   "86_Times_STEP_MAX_TIME_STP_350" : Time = PLC "86_Times".STEP_MAX_TIME_STP_350, 1 s
   "86_Times_STEP_MAX_TIME_STP_230" : Time = PLC "86_Times".STEP_MAX_TIME_STP_230, 1 s
   "20_TANKS_IP_DATA_RIO_02_FIRST_TANK_GTT_ISOL_VALVE_CLSD" : Bool = PLC "20_TANKS_IP_DATA".RIO_02.FIRST_TANK.GTT_ISOL_VALVE_CLSD AT %DB1.DBW0, 1 s
   "86_Times_STEP_MAX_TIME_STP_360" : Time = PLC "86_Times".STEP_MAX_TIME_STP_360, 1 s
   "40_TANKS_OP_DATA_RIO_02_VENT_B_2P" : Bool = PLC "40_TANKS_OP_DATA".RIO_02_VENT_B_2P AT %DB1.DBW0, 1 s
   "2019_AUT_MAN_CNTRL_STBD_GTT_VLV_MAN" : Bool = PLC "2019_AUT_MAN_CNTRL".STBD_GTT_VLV_MAN AT %DB1.DBW0, 1 s
   "14_DQ_DATA_CV_422_2P" : Bool = PLC "14_DQ_DATA".CV_422_2P AT %DB1.DBW0, 1 s
   "14_DQ_DATA_CV_421_2S" : Bool = PLC "14_DQ_DATA".CV_421_2S AT %DB1.DBW0, 1 s
   "2086_Times_DEOX_PRE_GTT_OPN_DLY" : Time = PLC "2086_Times".DEOX_PRE_GTT_OPN_DLY AT %DB1.DBW0, 1 s
   "2086_Times_DEOX_PRE_GTT_CLS_DLY" : Time = PLC "2086_Times".DEOX_PRE_GTT_CLS_DLY AT %DB1.DBW0, 1 s
   "2086_Times_REOX_PRE_GTT_OPN_DLY" : Time = PLC "2086_Times".REOX_PRE_GTT_OPN_DLY AT %DB1.DBW0, 1 s
   "2086_Times_REOX_PRE_GTT_CLS_DLY" : Time = PLC "2086_Times".REOX_PRE_GTT_CLS_DLY AT %DB1.DBW0, 1 s
   "2086_Times_AT_DEOX_CNF_TIME" : Time = PLC "2086_Times".AT_DEOX_CNF_TIME AT %DB1.DBW0, 1 s
   "2086_Times_AT_REOX_CNF_TIME" : Time = PLC "2086_Times".AT_REOX_CNF_TIME AT %DB1.DBW0, 1 s
   "2084_Setpoints_FIT418_LoLo" : Real = PLC "84_Setpoints".TIT401_High AT %DB1.DBW0, 1 s
   "2084_Setpoints_PIT424_HiHi" : Real = PLC "2084_Setpoints".PIT424_HiHi AT %DB1.DBW0, 1 s
   "2084_Setpoints_PIT424_Lo" : Real = PLC "2084_Setpoints".PIT424_Lo AT %DB1.DBW0, 1 s
   "2084_Setpoints_PIT424_LoLo" : Real = PLC "2084_Setpoints".PIT424_LoLo AT %DB1.DBW0, 1 s
   "2084_Setpoints_PIT415_HiHi" : Real = PLC "2084_Setpoints".PIT415_HiHi AT %DB1.DBW0, 1 s
   "2084_Setpoints_PIT415_Hi" : Real = PLC "2084_Setpoints".PIT415_Hi AT %DB1.DBW0, 1 s
   "2084_Setpoints_PIT415_Lo" : Real = PLC "2084_Setpoints".PIT415_Lo AT %DB1.DBW0, 1 s
   "2084_Setpoints_PIT415_LoLo" : Real = PLC "2084_Setpoints".PIT415_LoLo AT %DB1.DBW0, 1 s
   "2084_Setpoints_FIT418_Lo" : Real = PLC "2084_Setpoints".FIT418_Lo AT %DB1.DBW0, 1 s
   "2084_Setpoints_FIT418_Hi" : Real = PLC "2084_Setpoints".FIT418_Hi AT %DB1.DBW0, 1 s
   "20_TANKS_IP_DATA_RIO_02_FIRST_TANK_TANK_VENT_A_CLSD" : Bool = PLC "20_TANKS_IP_DATA".RIO_02.FIRST_TANK.TANK_VENT_A_CLSD AT %DB1.DBW0, 1 s
   "2084_Setpoints_TT436_HiHi" : Real = PLC "FIT418_FPT__ALM_ANALOG_DB"."VERY HIGH LEVEL VALUE (HH)" AT %DB1.DBW0, 1 s
   "2084_Setpoints_PH_SP" : Real = PLC "2084_Setpoints".PH_SP AT %DB1.DBW0, 1 s
   "2084_Setpoints_FIT418_HiHi" : Real = PLC "2084_Setpoints".FIT418_HiHi AT %DB1.DBW0, 1 s
   "2019_AUT_MAN_CNTRL_PORT_GTT_VLV_MAN" : Bool = PLC "2019_AUT_MAN_CNTRL".PORT_GTT_VLV_MAN AT %DB1.DBW0, 1 s
   "2084_Setpoints_FIT420_LoLo" : Real = PLC "2084_Setpoints".FIT420_LoLo AT %DB1.DBW0, 1 s
   "2084_Setpoints_FIT420_Hi" : Real = PLC "2084_Setpoints".FIT420_Hi AT %DB1.DBW0, 1 s
   "2084_Setpoints_FIT420_HiHi" : Real = PLC "2084_Setpoints".FIT420_HiHi AT %DB1.DBW0, 1 s
   "2084_Setpoints_LT422_Lo" : Real = PLC "2084_Setpoints".LT422_Lo AT %DB1.DBW0, 1 s
   "2084_Setpoints_LT422_Hi" : Real = PLC "2084_Setpoints".LT422_Hi AT %DB1.DBW0, 1 s
   "2084_Setpoints_TT436_Hi" : Real = PLC "2084_Setpoints".TT436_Hi AT %DB1.DBW0, 1 s
   "2084_Setpoints_DO_SP" : Real = PLC "2084_Setpoints".DO_SP AT %DB1.DBW0, 1 s
   "2084_Setpoints_FIT420_Lo" : Real = PLC "2084_Setpoints".FIT420_Lo AT %DB1.DBW0, 1 s
   "20_TANKS_IP_DATA_RIO_02_SECOND_TANK_GTT_ISOL_VALVE_CLSD" : Bool = PLC "20_TANKS_IP_DATA".RIO_02.SECOND_TANK.GTT_ISOL_VALVE_CLSD AT %DB1.DBW0, 1 s
   "2084_Setpoints_PIT424_Hi" : Real = PLC "2084_Setpoints".PIT424_Hi AT %DB1.DBW0, 1 s
   "20_TANKS_IP_DATA_RIO_02_SECOND_TANK_DECK_IG_PRESS" : Real = PLC "20_TANKS_IP_DATA".RIO_02.SECOND_TANK.DECK_IG_PRESS AT %DB1.DBW0, 1 s
   "20_TANKS_IP_DATA_RIO_02_FIRST_TANK_TANK_VENT_B_CLSD" : Bool = PLC "20_TANKS_IP_DATA".RIO_02.FIRST_TANK.TANK_VENT_B_CLSD AT %DB1.DBW0, 1 s
   "20_TANKS_IP_DATA_RIO_02_SECOND_TANK_GTT_ISOL_VALVE_OPEN" : Bool = PLC "20_TANKS_IP_DATA".RIO_02.SECOND_TANK.GTT_ISOL_VALVE_OPEN AT %DB1.DBW0, 1 s
   "20_TANKS_IP_DATA_RIO_02_FIRST_TANK_TANK_VENT_B_OPEN" : Bool = PLC "20_TANKS_IP_DATA".RIO_02.FIRST_TANK.TANK_VENT_B_OPEN AT %DB1.DBW0, 1 s
   "40_TANKS_OP_DATA_RIO_02_VENT_B_2P(1)" : Bool = PLC "40_TANKS_OP_DATA".RIO_02_VENT_B_2P AT %DB1.DBW0, 1 s
   "20_TANKS_IP_DATA_RIO_02_SECOND_TANK_TANK_VENT_B_CLSD" : Bool = PLC "20_TANKS_IP_DATA".RIO_02.SECOND_TANK.TANK_VENT_B_CLSD AT %DB1.DBW0, 1 s
   "40_TANKS_OP_DATA_RIO_02_VENT_B_2S(1)" : Bool = PLC "40_TANKS_OP_DATA".RIO_02_VENT_B_2S AT %DB1.DBW0, 1 s
   "20_TANKS_IP_DATA_RIO_02_SECOND_TANK_TANK_VENT_A_OPEN" : Bool = PLC "20_TANKS_IP_DATA".RIO_02.SECOND_TANK.TANK_VENT_A_OPEN AT %DB1.DBW0, 1 s
   "20_TANKS_IP_DATA_RIO_02_SECOND_TANK_TANK_VENT_A_CLSD" : Bool = PLC "20_TANKS_IP_DATA".RIO_02.SECOND_TANK.TANK_VENT_A_CLSD AT %DB1.DBW0, 1 s
   "20_TANKS_IP_DATA_RIO_02_FIRST_TANK_BWT_LEVEL_HIHI" : Bool = PLC "20_TANKS_IP_DATA".RIO_02.FIRST_TANK.BWT_LEVEL_HIHI AT %DB1.DBW0, 1 s
   "20_TANKS_IP_DATA_RIO_02_SECOND_TANK_BWT_LEVEL_HIHI" : Bool = PLC "20_TANKS_IP_DATA".RIO_02.SECOND_TANK.BWT_LEVEL_HIHI AT %DB1.DBW0, 1 s
   "20_TANKS_IP_DATA_RIO_02_SECOND_TANK_TANK_VENT_B_OPEN" : Bool = PLC "20_TANKS_IP_DATA".RIO_02.SECOND_TANK.TANK_VENT_B_OPEN AT %DB1.DBW0, 1 s
   "20_TANKS_IP_DATA_RIO_02_SECOND_TANK_TANKS_PRESS_HIHI" : Bool = PLC "20_TANKS_IP_DATA".RIO_02.SECOND_TANK.TANKS_PRESS_HIHI AT %DB1.DBW0, 1 s
   "20_TANKS_IP_DATA_RIO_02_SECOND_TANK_MBG_FLOW" : Real = PLC "20_TANKS_IP_DATA".RIO_02.SECOND_TANK.MBG_FLOW AT %DB1.DBW0, 1 s
   "20_TANKS_IP_DATA_RIO_02_FIRST_TANK_TANKS_PRESS" : Real = PLC "20_TANKS_IP_DATA".RIO_02.FIRST_TANK.TANKS_PRESS AT %DB1.DBW0, 1 s
   "20_TANKS_IP_DATA_RIO_02_FIRST_TANK_USD_FLOW" : Real = PLC "20_TANKS_IP_DATA".RIO_02.FIRST_TANK.USD_FLOW AT %DB1.DBW0, 1 s
   "20_TANKS_IP_DATA_RIO_02_FIRST_TANK_TANKS_PRESS_HIHI" : Bool = PLC "20_TANKS_IP_DATA".RIO_02.FIRST_TANK.TANKS_PRESS_HIHI AT %DB1.DBW0, 1 s
   "20_TANKS_IP_DATA_RIO_02_FIRST_TANK_MBG_FLOW" : Real = PLC "20_TANKS_IP_DATA".RIO_02.FIRST_TANK.MBG_FLOW AT %DB1.DBW0, 1 s
   "20_TANKS_IP_DATA_RIO_02_FIRST_TANK_O2_MONITOR" : Real = PLC "20_TANKS_IP_DATA".RIO_02.FIRST_TANK.O2_MONITOR AT %DB1.DBW0, 1 s
   "20_TANKS_IP_DATA_RIO_02_SECOND_TANK_USD_FLOW" : Real = PLC "20_TANKS_IP_DATA".RIO_02.SECOND_TANK.USD_FLOW AT %DB1.DBW0, 1 s
   "20_TANKS_IP_DATA_RIO_02_SECOND_TANK_TANKS_PRESS" : Real = PLC "20_TANKS_IP_DATA".RIO_02.SECOND_TANK.TANKS_PRESS AT %DB1.DBW0, 1 s
   "20_TANKS_IP_DATA_RIO_02_SECOND_TANK_O2_MONITOR" : Real = PLC "20_TANKS_IP_DATA".RIO_02.SECOND_TANK.O2_MONITOR AT %DB1.DBW0, 1 s
   "62_Warning_Data_GCU_WARNING_WORD_09(1)" : Word = PLC "62_Warning_Data".GCU_WARNING_WORD_09 AT %DB62.DBW16, 1 s
   "62_Warning_Data_GCU_WARNING_WORD_01(1)" : Word = PLC "62_Warning_Data".GCU_WARNING_WORD_01 AT %DB62.DBW0, 1 s
   "62_Warning_Data_BWTS_WARNING_WORD_10" : Word = PLC "62_Warning_Data".BWTS_WARNING_WORD_10 AT %DB62.DBW18, 1 s
   "62_Warning_Data_BWTS_WARNING_WORD_11" : Word = PLC "62_Warning_Data".BWTS_WARNING_WORD_11 AT %DB62.DBW20, 1 s
   "62_Warning_Data_GCU_WARNING_WORD_02(1)" : Word = PLC "62_Warning_Data".GCU_WARNING_WORD_02 AT %DB62.DBW2, 1 s
   "62_Warning_Data_GCU_WARNING_WORD_03(1)" : Word = PLC "62_Warning_Data".GCU_WARNING_WORD_03 AT %DB62.DBW4, 1 s
   "62_Warning_Data_GCU_WARNING_WORD_04(1)" : Word = PLC "62_Warning_Data".GCU_WARNING_WORD_04 AT %DB62.DBW6, 1 s
   "62_Warning_Data_GCU_WARNING_WORD_05(1)" : Word = PLC "62_Warning_Data".GCU_WARNING_WORD_05 AT %DB62.DBW8, 1 s
   "62_Warning_Data_GCU_WARNING_WORD_06(1)" : Word = PLC "62_Warning_Data".GCU_WARNING_WORD_06 AT %DB62.DBW10, 1 s
   "62_Warning_Data_GCU_WARNING_WORD_07(1)" : Word = PLC "62_Warning_Data".GCU_WARNING_WORD_07 AT %DB62.DBW12, 1 s
   "62_Warning_Data_GCU_WARNING_WORD_08(1)" : Word = PLC "62_Warning_Data".GCU_WARNING_WORD_08 AT %DB62.DBW14, 1 s
   "Record Data Tag" : Int AT %DB1.DBX0.0
   "Recipe Tag" : Int, internal
   "Data_From_WBT_Level_APT" : Real = PLC Data_From_WBT.Level_APT, 1 s
   "Data_From_WBT_Level_WBT_6P" : Real = PLC Data_From_WBT.Level_WBT_6P, 1 s
   "Data_From_WBT_Level_WBT_5P" : Real = PLC Data_From_WBT.Level_WBT_5P, 1 s
   "Data_From_WBT_Level_WBT_4P" : Real = PLC Data_From_WBT.Level_WBT_4P, 1 s
   "Data_From_WBT_Level_WBT_3P" : Real = PLC Data_From_WBT.Level_WBT_3P, 1 s
   "Data_From_WBT_Level_WBT_2P" : Real = PLC Data_From_WBT.Level_WBT_2P, 1 s
   "Data_From_WBT_Level_WBT_1P" : Real = PLC Data_From_WBT.Level_WBT_1P, 1 s
   "Data_From_WBT_Level_FPT" : Real = PLC Data_From_WBT.Level_FPT, 1 s
   "Data_From_WBT_Level_WBT_1S" : Real = PLC Data_From_WBT.Level_WBT_1S, 1 s
   "Data_From_WBT_Level_WBT_2S" : Real = PLC Data_From_WBT.Level_WBT_2S, 1 s
   "Data_From_WBT_Level_WBT_3S" : Real = PLC Data_From_WBT.Level_WBT_3S, 1 s
   "Data_From_WBT_Level_WBT_4S" : Real = PLC Data_From_WBT.Level_WBT_4S, 1 s
   "Data_From_WBT_Level_WBT_5S" : Real = PLC Data_From_WBT.Level_WBT_5S, 1 s
   "Data_From_WBT_Level_WBT_6S" : Real = PLC Data_From_WBT.Level_WBT_6S, 1 s
   "Data_From_WBT_Level_APT(1)" : Real = PLC Data_From_WBT.Level_APT, 1 s
   "Data_From_WBT_Level_APT m" : Real = PLC Data_From_WBT."Level_APT m", 1 s
   "Data_From_WBT_Level_WBT_6S m" : Real = PLC Data_From_WBT."Level_WBT_6S m", 1 s
   "Data_From_WBT_Level_WBT_5S m" : Real = PLC Data_From_WBT."Level_WBT_5S m", 1 s
   "Data_From_WBT_Level_WBT_4S m" : Real = PLC Data_From_WBT."Level_WBT_4S m", 1 s
   "Data_From_WBT_Level_WBT_3S m" : Real = PLC Data_From_WBT."Level_WBT_3S m", 1 s
   "Data_From_WBT_Level_WBT_2S m" : Real = PLC Data_From_WBT."Level_WBT_2S m", 1 s
   "Data_From_WBT_Level_WBT_1S m" : Real = PLC Data_From_WBT."Level_WBT_1S m", 1 s
   "Data_From_WBT_Level_FPT m" : Real = PLC Data_From_WBT."Level_FPT m", 1 s
   "Data_From_WBT_Level_WBT_1P m" : Real = PLC Data_From_WBT."Level_WBT_1P m", 1 s
   "Data_From_WBT_Level_WBT_2P m" : Real = PLC Data_From_WBT."Level_WBT_2P m", 1 s
   "Data_From_WBT_Level_WBT_3P m" : Real = PLC Data_From_WBT."Level_WBT_3P m", 1 s
   "Data_From_WBT_Level_WBT_4P m" : Real = PLC Data_From_WBT."Level_WBT_4P m", 1 s
   "Data_From_WBT_Level_WBT_5P m" : Real = PLC Data_From_WBT."Level_WBT_5P m", 1 s
   "Data_From_WBT_Level_WBT_6P m" : Real = PLC Data_From_WBT."Level_WBT_6P m", 1 s
   "HEART BEAT TRUE" : Bool = PLC "68_Sys_Status_Data"."TRUE for HMI" AT %M1.2, 100 ms
   "Warn To Start IGG" : Bool = PLC "82_To_HMI"."Warn to Start IGG", 1 s
      on ChangeValue: "TimeRemainingToTreatment"()

discrete alarms
   129: 'PIT-359 - HIGH HIGH', class IGG Alarms, trigger "Alarms_Acknowledge_IGG_ALARM_ACKNLG_2" bit 1
   130: 'PIT-316 - HIGH HIGH', class IGG Alarms, trigger "Alarms_Acknowledge_IGG_ALARM_ACKNLG_2" bit 3
   131: 'PIT-359 - LOW LOW', class IGG Alarms, trigger "Alarms_Acknowledge_IGG_ALARM_ACKNLG_2" bit 0
   132: 'PIT-316 - LOW LOW', class IGG Alarms, trigger "Alarms_Acknowledge_IGG_ALARM_ACKNLG_2" bit 2
   279: 'IGG_MESSAGE_WORD_02_BIT_14', class IGG Messages, trigger "64_Message_Data_IGG_MESSAGE_WORD_02" bit 6
   133: 'PIT-359 - HIGH HIGH', class IGG Alarms, trigger "Alarms_Acknowledge_IGG_ALARM_ACKNLG_2" bit 4
   134: 'TIT-401 - HIGH HIGH', class IGG Alarms, trigger "Alarms_Acknowledge_IGG_ALARM_ACKNLG_2" bit 10
   135: 'PIT-102 CA PRESSURE - FAULT', class IGG Alarms, trigger "Alarms_Acknowledge_IGG_ALARM_ACKNLG_2" bit 9
   136: 'PIT-402 IG OUTLET PRESSURE - HIGH HIGH', class IGG Alarms, trigger "Alarms_Acknowledge_IGG_ALARM_ACKNLG_2" bit 12
   137: 'PIT-402 IG OUTLET PRESSURE - LOW LOW', class IGG Alarms, trigger "Alarms_Acknowledge_IGG_ALARM_ACKNLG_2" bit 11
   138: 'IGG_ALARM_WORD_02_BIT_14', class IGG Alarms, trigger "Alarms_Acknowledge_IGG_ALARM_ACKNLG_2" bit 6
   139: 'IGG_ALARM_WORD_02_BIT_13', class IGG Alarms, trigger "Alarms_Acknowledge_IGG_ALARM_ACKNLG_2" bit 5
   140: 'PIT-102 CA PRESSURE - LOW LOW', class IGG Alarms, trigger "Alarms_Acknowledge_IGG_ALARM_ACKNLG_2" bit 8
   141: 'IGG_ALARM_WORD_02_BIT_15', class IGG Alarms, trigger "Alarms_Acknowledge_IGG_ALARM_ACKNLG_2" bit 7
   142: 'EMERGENCY STOP ACTIVE', class IGG Alarms, trigger "Alarms_Acknowledge_IGG_ALARM_ACKNLG_1" bit 15
   143: 'ATMOSPHERIC O2 SENSOR 1 - LOW LOW', class IGG Alarms, trigger "Alarms_Acknowledge_IGG_ALARM_ACKNLG_1" bit 1
   144: 'BC ALARM ACTIVE', class IGG Alarms, trigger "Alarms_Acknowledge_IGG_ALARM_ACKNLG_1" bit 0
   145: 'ATMOSPHERIC O2 SENSOR 2 - LOW LOW', class IGG Alarms, trigger "Alarms_Acknowledge_IGG_ALARM_ACKNLG_1" bit 2
   146: 'E-500B FUEL PUMP - NOT RUNNING', class IGG Alarms, trigger "Alarms_Acknowledge_IGG_ALARM_ACKNLG_1" bit 4
   147: 'E-500A FUEL PUMP - NOT RUNNING', class IGG Alarms, trigger "Alarms_Acknowledge_IGG_ALARM_ACKNLG_1" bit 3
   383: 'BC_EVENT_WORD_02_BIT_6', class BC Events, trigger "66_Event_Data_BC_EVENT_WORD_02" bit 14
   382: 'BC_EVENT_WORD_02_BIT_5', class BC Events, trigger "66_Event_Data_BC_EVENT_WORD_02" bit 13
   384: 'BC_EVENT_WORD_02_BIT_7', class BC Events, trigger "66_Event_Data_BC_EVENT_WORD_02" bit 15
   278: 'IGG_MESSAGE_WORD_02_BIT_13', class IGG Messages, trigger "64_Message_Data_IGG_MESSAGE_WORD_02" bit 5
   277: 'IGG_MESSAGE_WORD_02_BIT_12', class IGG Messages, trigger "64_Message_Data_IGG_MESSAGE_WORD_02" bit 4
   148: 'P-301 CSW PUMP - TRIPPED', class IGG Alarms, trigger "Alarms_Acknowledge_IGG_ALARM_ACKNLG_1" bit 11
   149: 'IGG AUTO INTERLOCKS NOT OK', class IGG Alarms, trigger "Alarms_Acknowledge_IGG_ALARM_ACKNLG_1" bit 10
   150: 'E-500A FUEL PUMP - TRIPPED', class IGG Alarms, trigger "Alarms_Acknowledge_IGG_ALARM_ACKNLG_1" bit 12
   151: 'E-139 CAB INVERTER - FAULT', class IGG Alarms, trigger "Alarms_Acknowledge_IGG_ALARM_ACKNLG_1" bit 14
   152: 'E-500B FUEL PUMP - TRIPPED', class IGG Alarms, trigger "Alarms_Acknowledge_IGG_ALARM_ACKNLG_1" bit 13
   153: 'IGG_ALARM_WORD_01_BIT_14', class IGG Alarms, trigger "Alarms_Acknowledge_IGG_ALARM_ACKNLG_1" bit 6
   154: 'E-139 CAB NOT READY3', class IGG Alarms, trigger "Alarms_Acknowledge_IGG_ALARM_ACKNLG_1" bit 5
   155: 'IGG_ALARM_WORD_01_BIT_15', class IGG Alarms, trigger "Alarms_Acknowledge_IGG_ALARM_ACKNLG_1" bit 7
   156: 'SLAVE PLC HEART BEAT MISSING', class IGG Alarms, trigger "Alarms_Acknowledge_IGG_ALARM_ACKNLG_1" bit 9
   157: 'MASTER PLC HEART BEAT MISSING', class IGG Alarms, trigger "Alarms_Acknowledge_IGG_ALARM_ACKNLG_1" bit 8
   158: 'PIT-402 IG PRESSURE - OUT OF RANGE', class IGG Alarms, trigger "Alarms_Acknowledge_IGG_ALARM_ACKNLG_2" bit 13
   55: 'IGG_ALARM_WORD_04_BIT_14', class IGG Alarms, trigger "Alarms_Acknowledge_IGG_ALARM_ACKNLG_4" bit 6
   54: 'CORRECT PHASE ROTATION - FAULT', class IGG Alarms, trigger "Alarms_Acknowledge_IGG_ALARM_ACKNLG_4" bit 5
   56: 'IGG_ALARM_WORD_04_BIT_15', class IGG Alarms, trigger "Alarms_Acknowledge_IGG_ALARM_ACKNLG_4" bit 7
   58: 'CV-312 - FAULT', class IGG Alarms, trigger "Alarms_Acknowledge_IGG_ALARM_ACKNLG_4" bit 9
   57: 'CV-311 - FAULT', class IGG Alarms, trigger "Alarms_Acknowledge_IGG_ALARM_ACKNLG_4" bit 8
   50: 'TIT-319 INLET CSW TEMP - FAULT AND TIT-401 AND TIT-360 - FAULT', class IGG Alarms, trigger "Alarms_Acknowledge_IGG_ALARM_ACKNLG_4" bit 1
   49: 'TIT-319 INLET CSW TEMP - FAULT AND TS-006 - FAULT', class IGG Alarms, trigger "Alarms_Acknowledge_IGG_ALARM_ACKNLG_4" bit 0
   51: 'TIT-360 OUTLET CSW TEMP - HIGH HIGH0', class IGG Alarms, trigger "Alarms_Acknowledge_IGG_ALARM_ACKNLG_4" bit 2
   53: 'E-139 NOT RUNNING2', class IGG Alarms, trigger "Alarms_Acknowledge_IGG_ALARM_ACKNLG_4" bit 4
   52: 'TIT-360 OUTLET CSW TEMP - HIGH HIGH AND TIT-401 - FAULT', class IGG Alarms, trigger "Alarms_Acknowledge_IGG_ALARM_ACKNLG_4" bit 3
   59: 'CV-321 - FAULT', class IGG Alarms, trigger "Alarms_Acknowledge_IGG_ALARM_ACKNLG_4" bit 10
   65: 'IGG ALARM ACTIVE', class BC Alarms, trigger "BC_ALARM_ACKNLG_1" bit 0
   282: 'IGG_MESSAGE_WORD_02_BIT_1', class IGG Messages, trigger "64_Message_Data_IGG_MESSAGE_WORD_02" bit 9
   66: 'PS-101 PRESSURE NOT PRESENT - FAULT', class BC Alarms, trigger "BC_ALARM_ACKNLG_1" bit 1
   69: 'FD-001 FLAME SIGNAL - OUT OF RANGE', class BC Alarms, trigger "BC_ALARM_ACKNLG_1" bit 4
   68: 'O2 SYSTEM POWER NOT HEALTHY', class BC Alarms, trigger "BC_ALARM_ACKNLG_1" bit 3
   61: 'CV-401 - FAULT', class IGG Alarms, trigger "Alarms_Acknowledge_IGG_ALARM_ACKNLG_4" bit 12
   60: 'CV-322 - FAULT', class IGG Alarms, trigger "Alarms_Acknowledge_IGG_ALARM_ACKNLG_4" bit 11
   62: 'CV-431 - FAULT', class IGG Alarms, trigger "Alarms_Acknowledge_IGG_ALARM_ACKNLG_4" bit 13
   64: 'SAFETY SYSTEM INTERLOCK', class IGG Alarms, trigger "Alarms_Acknowledge_IGG_ALARM_ACKNLG_4" bit 15
   63: 'CV-432 - FAULT', class IGG Alarms, trigger "Alarms_Acknowledge_IGG_ALARM_ACKNLG_4" bit 14
   35: 'TIT-315 SHELL CSW TEMP - HIGH HIGH AND TIT-401 - FAULT', class IGG Alarms, trigger "Alarms_Acknowledge_IGG_ALARM_ACKNLG_3" bit 2
   34: 'TIT-315 SHELL CSW TEMP - HIGH HIGH AND TS-006 - FAULT', class IGG Alarms, trigger "Alarms_Acknowledge_IGG_ALARM_ACKNLG_3" bit 1
   36: 'PIT-316 OUTLET CSW PRESSURE AND FS-317 - FAULT', class IGG Alarms, trigger "Alarms_Acknowledge_IGG_ALARM_ACKNLG_3" bit 3
   38: 'PIT-316 OUTLET CSW PRESSURE AND TS-006 - FAULT', class IGG Alarms, trigger "Alarms_Acknowledge_IGG_ALARM_ACKNLG_3" bit 5
   37: 'PIT-316 OUTLET CSW PRESSURE AND TIT-315 - FAULT', class IGG Alarms, trigger "Alarms_Acknowledge_IGG_ALARM_ACKNLG_3" bit 4
   159: 'TIT-360 - HIGH HIGH', class IGG Alarms, trigger "Alarms_Acknowledge_IGG_ALARM_ACKNLG_2" bit 15
   160: 'TIT-319 - HIGH HIGH', class IGG Alarms, trigger "Alarms_Acknowledge_IGG_ALARM_ACKNLG_2" bit 14
   280: 'IGG_MESSAGE_WORD_02_BIT_15', class IGG Messages, trigger "64_Message_Data_IGG_MESSAGE_WORD_02" bit 7
   33: 'TIT-315 SHELL CSW TEMP - HIGH HIGH AND FS-317 - FAULT', class IGG Alarms, trigger "Alarms_Acknowledge_IGG_ALARM_ACKNLG_3" bit 0
   70: 'E-600 O2 ANALYSER CONTENT - OUT OF RANGE', class BC Alarms, trigger "BC_ALARM_ACKNLG_1" bit 5
   39: 'IGG_ALARM_WORD_03_BIT_14', class IGG Alarms, trigger "Alarms_Acknowledge_IGG_ALARM_ACKNLG_3" bit 6
   46: 'TIT-401 IG TEMP - HIGH HIGH AND TIT-360 - FAULT', class IGG Alarms, trigger "Alarms_Acknowledge_IGG_ALARM_ACKNLG_3" bit 13
   45: 'TIT-401 IG TEMP - HIGH HIGH AND TS-403 - FAULT', class IGG Alarms, trigger "Alarms_Acknowledge_IGG_ALARM_ACKNLG_3" bit 12
   47: 'IGG_ALARM_WORD_03_BIT_6', class IGG Alarms, trigger "Alarms_Acknowledge_IGG_ALARM_ACKNLG_3" bit 14
   281: 'IGG_MESSAGE_WORD_02_BIT_0', class IGG Messages, trigger "64_Message_Data_IGG_MESSAGE_WORD_02" bit 8
   48: 'IGG_ALARM_WORD_03_BIT_7', class IGG Alarms, trigger "Alarms_Acknowledge_IGG_ALARM_ACKNLG_3" bit 15
   41: 'PIT-112/113 TIER ALARM - PRESSURE NOT OK', class IGG Alarms, trigger "Alarms_Acknowledge_IGG_ALARM_ACKNLG_3" bit 8
   40: 'IGG_ALARM_WORD_03_BIT_15', class IGG Alarms, trigger "Alarms_Acknowledge_IGG_ALARM_ACKNLG_3" bit 7
   42: 'PIT-102 CA PRESSURE - LOW LOW AND FDU - FAULT', class IGG Alarms, trigger "Alarms_Acknowledge_IGG_ALARM_ACKNLG_3" bit 9
   44: 'IGG ALARM WORD', class IGG Alarms, trigger "Alarms_Acknowledge_IGG_ALARM_ACKNLG_3" bit 11
   43: 'PIT-102 CA PRESSURE - LOW LOW AND PIT-402 - FAULT', class IGG Alarms, trigger "Alarms_Acknowledge_IGG_ALARM_ACKNLG_3" bit 10
   381: 'BC_EVENT_WORD_02_BIT_4', class BC Events, trigger "66_Event_Data_BC_EVENT_WORD_02" bit 12
   330: 'IGG_EVENT_WORD_01_BIT_1', class IGG Events, trigger "66_Event_Data_IGG_EVENT_WORD_01" bit 9
   329: 'IGG_EVENT_WORD_01_BIT_0', class IGG Events, trigger "66_Event_Data_IGG_EVENT_WORD_01" bit 8
   331: 'IGG_EVENT_WORD_01_BIT_2', class IGG Events, trigger "66_Event_Data_IGG_EVENT_WORD_01" bit 10
   333: 'IGG_EVENT_WORD_01_BIT_4', class IGG Events, trigger "66_Event_Data_IGG_EVENT_WORD_01" bit 12
   332: 'IGG_EVENT_WORD_01_BIT_3', class IGG Events, trigger "66_Event_Data_IGG_EVENT_WORD_01" bit 11
   325: 'IGG_EVENT_WORD_01_BIT_12', class IGG Events, trigger "66_Event_Data_IGG_EVENT_WORD_01" bit 4
   324: 'IGG_EVENT_WORD_01_BIT_11', class IGG Events, trigger "66_Event_Data_IGG_EVENT_WORD_01" bit 3
   326: 'IGG_EVENT_WORD_01_BIT_13', class IGG Events, trigger "66_Event_Data_IGG_EVENT_WORD_01" bit 5
   328: 'IGG_EVENT_WORD_01_BIT_15', class IGG Events, trigger "66_Event_Data_IGG_EVENT_WORD_01" bit 7
   327: 'IGG_EVENT_WORD_01_BIT_14', class IGG Events, trigger "66_Event_Data_IGG_EVENT_WORD_01" bit 6
   338: 'IGG_EVENT_WORD_02_BIT_9', class IGG Events, trigger "66_Event_Data_IGG_EVENT_WORD_02" bit 1
   337: 'IGG_EVENT_WORD_02_BIT_8', class IGG Events, trigger "66_Event_Data_IGG_EVENT_WORD_02" bit 0
   339: 'IGG_EVENT_WORD_02_BIT_10', class IGG Events, trigger "66_Event_Data_IGG_EVENT_WORD_02" bit 2
   341: 'IGG_EVENT_WORD_02_BIT_12', class IGG Events, trigger "66_Event_Data_IGG_EVENT_WORD_02" bit 4
   340: 'IGG_EVENT_WORD_02_BIT_11', class IGG Events, trigger "66_Event_Data_IGG_EVENT_WORD_02" bit 3
   335: 'IGG_EVENT_WORD_01_BIT_6', class IGG Events, trigger "66_Event_Data_IGG_EVENT_WORD_01" bit 14
   334: 'IGG_EVENT_WORD_01_BIT_5', class IGG Events, trigger "66_Event_Data_IGG_EVENT_WORD_01" bit 13
   336: 'IGG_EVENT_WORD_01_BIT_7', class IGG Events, trigger "66_Event_Data_IGG_EVENT_WORD_01" bit 15
   276: 'IGG_MESSAGE_WORD_02_BIT_11', class IGG Messages, trigger "64_Message_Data_IGG_MESSAGE_WORD_02" bit 3
   259: 'IGG_MESSAGE_WORD_01_BIT_10', class IGG Messages, trigger "64_Message_Data_IGG_MESSAGE_WORD_01" bit 2
   267: 'IGG_MESSAGE_WORD_01_BIT_2', class IGG Messages, trigger "64_Message_Data_IGG_MESSAGE_WORD_01" bit 10
   268: 'IGG_MESSAGE_WORD_01_BIT_3', class IGG Messages, trigger "64_Message_Data_IGG_MESSAGE_WORD_01" bit 11
   273: 'IGG_MESSAGE_WORD_02_BIT_8', class IGG Messages, trigger "64_Message_Data_IGG_MESSAGE_WORD_02" bit 0
   265: 'IGG_MESSAGE_WORD_01_BIT_0', class IGG Messages, trigger "64_Message_Data_IGG_MESSAGE_WORD_01" bit 8
   266: 'IGG_MESSAGE_WORD_01_BIT_1', class IGG Messages, trigger "64_Message_Data_IGG_MESSAGE_WORD_01" bit 9
   272: 'IGG_MESSAGE_WORD_01_BIT_7', class IGG Messages, trigger "64_Message_Data_IGG_MESSAGE_WORD_01" bit 15
   67: 'E-600 O2 ANALYSER SYSTEM - FAIL', class BC Alarms, trigger "BC_ALARM_ACKNLG_1" bit 2
   271: 'IGG_MESSAGE_WORD_01_BIT_6', class IGG Messages, trigger "64_Message_Data_IGG_MESSAGE_WORD_01" bit 14
   269: 'IGG_MESSAGE_WORD_01_BIT_4', class IGG Messages, trigger "64_Message_Data_IGG_MESSAGE_WORD_01" bit 12
   270: 'IGG_MESSAGE_WORD_01_BIT_5', class IGG Messages, trigger "64_Message_Data_IGG_MESSAGE_WORD_01" bit 13
   260: 'IGG_MESSAGE_WORD_01_BIT_11', class IGG Messages, trigger "64_Message_Data_IGG_MESSAGE_WORD_01" bit 3
   275: 'IGG_MESSAGE_WORD_02_BIT_10', class IGG Messages, trigger "64_Message_Data_IGG_MESSAGE_WORD_02" bit 2
   321: 'IGG_EVENT_WORD_01_BIT_8', class IGG Events, trigger "66_Event_Data_IGG_EVENT_WORD_01" bit 0
   323: 'IGG_EVENT_WORD_01_BIT_10', class IGG Events, trigger "66_Event_Data_IGG_EVENT_WORD_01" bit 2
   322: 'IGG_EVENT_WORD_01_BIT_9', class IGG Events, trigger "66_Event_Data_IGG_EVENT_WORD_01" bit 1
   264: 'IGG_MESSAGE_WORD_01_BIT_15', class IGG Messages, trigger "64_Message_Data_IGG_MESSAGE_WORD_01" bit 7
   274: 'IGG_MESSAGE_WORD_02_BIT_9', class IGG Messages, trigger "64_Message_Data_IGG_MESSAGE_WORD_02" bit 1
   263: 'IGG_MESSAGE_WORD_01_BIT_14', class IGG Messages, trigger "64_Message_Data_IGG_MESSAGE_WORD_01" bit 6
   261: 'IGG_MESSAGE_WORD_01_BIT_12', class IGG Messages, trigger "64_Message_Data_IGG_MESSAGE_WORD_01" bit 4
   262: 'IGG_MESSAGE_WORD_01_BIT_13', class IGG Messages, trigger "64_Message_Data_IGG_MESSAGE_WORD_01" bit 5
   342: 'IGG_EVENT_WORD_02_BIT_13', class IGG Events, trigger "66_Event_Data_IGG_EVENT_WORD_02" bit 5
   367: 'BC_EVENT_WORD_01_BIT_6', class BC Events, trigger "66_Event_Data_BC_EVENT_WORD_01" bit 14
   366: 'BC_EVENT_WORD_01_BIT_5', class BC Events, trigger "66_Event_Data_BC_EVENT_WORD_01" bit 13
   368: 'BC_EVENT_WORD_01_BIT_7', class BC Events, trigger "66_Event_Data_BC_EVENT_WORD_01" bit 15
   370: 'BC_EVENT_WORD_02_BIT_9', class BC Events, trigger "66_Event_Data_BC_EVENT_WORD_02" bit 1
   369: 'BC_EVENT_WORD_02_BIT_8', class BC Events, trigger "66_Event_Data_BC_EVENT_WORD_02" bit 0
   362: 'BC_EVENT_WORD_01_BIT_1', class BC Events, trigger "66_Event_Data_BC_EVENT_WORD_01" bit 9
   361: 'BC_EVENT_WORD_01_BIT_0', class BC Events, trigger "66_Event_Data_BC_EVENT_WORD_01" bit 8
   363: 'BC_EVENT_WORD_01_BIT_2', class BC Events, trigger "66_Event_Data_BC_EVENT_WORD_01" bit 10
   365: 'BC_EVENT_WORD_01_BIT_4', class BC Events, trigger "66_Event_Data_BC_EVENT_WORD_01" bit 12
   364: 'BC_EVENT_WORD_01_BIT_3', class BC Events, trigger "66_Event_Data_BC_EVENT_WORD_01" bit 11
   377: 'BC_EVENT_WORD_02_BIT_0', class BC Events, trigger "66_Event_Data_BC_EVENT_WORD_02" bit 8
   376: 'BC_EVENT_WORD_02_BIT_15', class BC Events, trigger "66_Event_Data_BC_EVENT_WORD_02" bit 7
   378: 'BC_EVENT_WORD_02_BIT_1', class BC Events, trigger "66_Event_Data_BC_EVENT_WORD_02" bit 9
   380: 'BC_EVENT_WORD_02_BIT_3', class BC Events, trigger "66_Event_Data_BC_EVENT_WORD_02" bit 11
   379: 'BC_EVENT_WORD_02_BIT_2', class BC Events, trigger "66_Event_Data_BC_EVENT_WORD_02" bit 10
   372: 'BC_EVENT_WORD_02_BIT_11', class BC Events, trigger "66_Event_Data_BC_EVENT_WORD_02" bit 3
   371: 'BC_EVENT_WORD_02_BIT_10', class BC Events, trigger "66_Event_Data_BC_EVENT_WORD_02" bit 2
   373: 'BC_EVENT_WORD_02_BIT_12', class BC Events, trigger "66_Event_Data_BC_EVENT_WORD_02" bit 4
   375: 'BC_EVENT_WORD_02_BIT_14', class BC Events, trigger "66_Event_Data_BC_EVENT_WORD_02" bit 6
   374: 'BC_EVENT_WORD_02_BIT_13', class BC Events, trigger "66_Event_Data_BC_EVENT_WORD_02" bit 5
   349: 'IGG_EVENT_WORD_02_BIT_4', class IGG Events, trigger "66_Event_Data_IGG_EVENT_WORD_02" bit 12
   348: 'IGG_EVENT_WORD_02_BIT_3', class IGG Events, trigger "66_Event_Data_IGG_EVENT_WORD_02" bit 11
   350: 'IGG_EVENT_WORD_02_BIT_5', class IGG Events, trigger "66_Event_Data_IGG_EVENT_WORD_02" bit 13
   352: 'IGG_EVENT_WORD_02_BIT_7', class IGG Events, trigger "66_Event_Data_IGG_EVENT_WORD_02" bit 15
   351: 'IGG_EVENT_WORD_02_BIT_6', class IGG Events, trigger "66_Event_Data_IGG_EVENT_WORD_02" bit 14
   344: 'IGG_EVENT_WORD_02_BIT_15', class IGG Events, trigger "66_Event_Data_IGG_EVENT_WORD_02" bit 7
   343: 'IGG_EVENT_WORD_02_BIT_14', class IGG Events, trigger "66_Event_Data_IGG_EVENT_WORD_02" bit 6
   345: 'IGG_EVENT_WORD_02_BIT_0', class IGG Events, trigger "66_Event_Data_IGG_EVENT_WORD_02" bit 8
   347: 'IGG_EVENT_WORD_02_BIT_2', class IGG Events, trigger "66_Event_Data_IGG_EVENT_WORD_02" bit 10
   346: 'IGG_EVENT_WORD_02_BIT_1', class IGG Events, trigger "66_Event_Data_IGG_EVENT_WORD_02" bit 9
   357: 'BC_EVENT_WORD_01_BIT_12', class BC Events, trigger "66_Event_Data_BC_EVENT_WORD_01" bit 4
   356: 'BC_EVENT_WORD_01_BIT_11', class BC Events, trigger "66_Event_Data_BC_EVENT_WORD_01" bit 3
   358: 'BC_EVENT_WORD_01_BIT_13', class BC Events, trigger "66_Event_Data_BC_EVENT_WORD_01" bit 5
   360: 'BC_EVENT_WORD_01_BIT_15', class BC Events, trigger "66_Event_Data_BC_EVENT_WORD_01" bit 7
   359: 'BC_EVENT_WORD_01_BIT_14', class BC Events, trigger "66_Event_Data_BC_EVENT_WORD_01" bit 6
   257: 'IGG_MESSAGE_WORD_01_BIT_8', class IGG Messages, trigger "64_Message_Data_IGG_MESSAGE_WORD_01" bit 0
   258: 'IGG_MESSAGE_WORD_01_BIT_9', class IGG Messages, trigger "64_Message_Data_IGG_MESSAGE_WORD_01" bit 1
   353: 'BC_EVENT_WORD_01_BIT_8', class BC Events, trigger "66_Event_Data_BC_EVENT_WORD_01" bit 0
   355: 'BC_EVENT_WORD_01_BIT_10', class BC Events, trigger "66_Event_Data_BC_EVENT_WORD_01" bit 2
   354: 'BC_EVENT_WORD_01_BIT_9', class BC Events, trigger "66_Event_Data_BC_EVENT_WORD_01" bit 1
   114: 'P-305 FRESH WATER PUMP - TRIPPED', class BC Alarms, trigger "BC_ALARM_ACKNLG_4" bit 1
   113: 'LS-001 IGG QUENCH CHAMBER LEVEL - HIGH', class BC Alarms, trigger "BC_ALARM_ACKNLG_4" bit 0
   116: 'BC_ALARM_WORD_04_BIT_11', class BC Alarms, trigger "BC_ALARM_ACKNLG_4" bit 3
   115: 'BC_ALARM_WORD_04_BIT_10', class BC Alarms, trigger "BC_ALARM_ACKNLG_4" bit 2
   284: 'IGG_MESSAGE_WORD_02_BIT_3', class IGG Messages, trigger "64_Message_Data_IGG_MESSAGE_WORD_02" bit 11
   112: 'BC_ALARM_WORD_3_BIT_15', class BC Alarms, trigger "BC_ALARM_ACKNLG_3" bit 15
   315: 'BC_MESSAGE_WORD_02_BIT_2', class BC Messages, trigger "64_Message_Data_BC_MESSAGE_WORD_02" bit 10
   316: 'BC_MESSAGE_WORD_02_BIT_3', class BC Messages, trigger "64_Message_Data_BC_MESSAGE_WORD_02" bit 11
   122: 'TS-006 IG SHELL TEMP HI SWITCH AND TIT-360 - FAULT', class BC Alarms, trigger "BC_ALARM_ACKNLG_4" bit 9
   121: 'TS-006 IGG SHELL TEMPERATURE - HIGH', class BC Alarms, trigger "BC_ALARM_ACKNLG_4" bit 8
   124: 'TS-403 IG TEMP - HIGH HIGH SWITCH AND TIT-401 - FAULT', class BC Alarms, trigger "BC_ALARM_ACKNLG_4" bit 11
   123: 'TS-006 IG SHELL TEMP HI SWITCH AND TIT-401 - FAULT', class BC Alarms, trigger "BC_ALARM_ACKNLG_4" bit 10
   297: 'BC_MESSAGE_WORD_01_BIT_0', class BC Messages, trigger "64_Message_Data_BC_MESSAGE_WORD_01" bit 8
   117: 'BC_ALARM_WORD_04_BIT_12', class BC Alarms, trigger "BC_ALARM_ACKNLG_4" bit 4
   120: 'BC_ALARM_WORD_04_BIT_15', class BC Alarms, trigger "BC_ALARM_ACKNLG_4" bit 7
   119: 'BC_ALARM_WORD_04_BIT_14', class BC Alarms, trigger "BC_ALARM_ACKNLG_4" bit 6
   111: 'BC_ALARM_WORD_03_BIT_6', class BC Alarms, trigger "BC_ALARM_ACKNLG_3" bit 14
   100: 'FS-317 JACKET COOLING WATER FLOW SWITCH - FAULT AND FS-320 - FAULT AND PIT 360 - FAULT', class BC Alarms, trigger "BC_ALARM_ACKNLG_3" bit 3
   99: 'FS-320 COOLING WATER FLOW SWITCH - FAULT AND TIT-401 - FAULT0', class BC Alarms, trigger "BC_ALARM_ACKNLG_3" bit 2
   102: 'FS-317 JACKET COOLING WATER FLOW SWITCH - FAULT AND TIT-401 - FAULT', class BC Alarms, trigger "BC_ALARM_ACKNLG_3" bit 5
   101: 'FS-317 JACKET COOLING WATER FLOW SWITCH FASULT AND TIT-360 - FAULT', class BC Alarms, trigger "BC_ALARM_ACKNLG_3" bit 4
   317: 'BC_MESSAGE_WORD_02_BIT_4', class BC Messages, trigger "64_Message_Data_BC_MESSAGE_WORD_02" bit 12
   318: 'BC_MESSAGE_WORD_02_BIT_5', class BC Messages, trigger "64_Message_Data_BC_MESSAGE_WORD_02" bit 13
   98: 'FS-320 COOLING WATER FLOW SWITCH - FAULT AND TIT-360 - FAULT', class BC Alarms, trigger "BC_ALARM_ACKNLG_3" bit 1
   97: 'FS-320 COOLING WATER FLOW SWITCH - FAULT AND FS-317 - FAULT', class BC Alarms, trigger "BC_ALARM_ACKNLG_3" bit 0
   108: 'PIT-112 INSTRUMENT AIR PRESSURE - FAULT AND FS-115 - FAULT', class BC Alarms, trigger "BC_ALARM_ACKNLG_3" bit 11
   107: 'PIT-112 INSTRUMENT AIR PRESSURE - FAULT', class BC Alarms, trigger "BC_ALARM_ACKNLG_3" bit 10
   110: 'FS-115 MAIN BURNER ATOMISING AIR FLOW SWITCH - FAULT AND PIT-113 - FAULT', class BC Alarms, trigger "BC_ALARM_ACKNLG_3" bit 13
   109: 'FS-115 MAIN BURNER ATOMISING AIR FLOW SWITCH - FAULT AND CV 114 CLOSE', class BC Alarms, trigger "BC_ALARM_ACKNLG_3" bit 12
   104: 'TS-403 IG VENT TEMPERATURE HIGH', class BC Alarms, trigger "BC_ALARM_ACKNLG_3" bit 7
   103: 'BC_ALARM_WORD_03_BIT_14', class BC Alarms, trigger "BC_ALARM_ACKNLG_3" bit 6
   106: 'FS-123 PILOT BURNER AIR FLOW SWITCH - FAULT AND PIT-112 LOW LOW', class BC Alarms, trigger "BC_ALARM_ACKNLG_3" bit 9
   105: 'FS-123 PILOT BURNER AIR FLOW SWITCH - FAULT AND PIT-112 HIGH HIGH', class BC Alarms, trigger "BC_ALARM_ACKNLG_3" bit 8
   305: 'BC_MESSAGE_WORD_02_BIT_8', class BC Messages, trigger "64_Message_Data_BC_MESSAGE_WORD_02" bit 0
   306: 'BC_MESSAGE_WORD_02_BIT_9', class BC Messages, trigger "64_Message_Data_BC_MESSAGE_WORD_02" bit 1
   304: 'BC_MESSAGE_WORD_01_BIT_7', class BC Messages, trigger "64_Message_Data_BC_MESSAGE_WORD_01" bit 15
   294: 'BC_MESSAGE_WORD_01_BIT_13', class BC Messages, trigger "64_Message_Data_BC_MESSAGE_WORD_01" bit 5
   293: 'BC_MESSAGE_WORD_01_BIT_12', class BC Messages, trigger "64_Message_Data_BC_MESSAGE_WORD_01" bit 4
   309: 'BC_MESSAGE_WORD_02_BIT_12', class BC Messages, trigger "64_Message_Data_BC_MESSAGE_WORD_02" bit 4
   307: 'BC_MESSAGE_WORD_02_BIT_10', class BC Messages, trigger "64_Message_Data_BC_MESSAGE_WORD_02" bit 2
   308: 'BC_MESSAGE_WORD_02_BIT_11', class BC Messages, trigger "64_Message_Data_BC_MESSAGE_WORD_02" bit 3
   300: 'BC_MESSAGE_WORD_01_BIT_3', class BC Messages, trigger "64_Message_Data_BC_MESSAGE_WORD_01" bit 11
   296: 'BC_MESSAGE_WORD_01_BIT_15', class BC Messages, trigger "64_Message_Data_BC_MESSAGE_WORD_01" bit 7
   298: 'BC_MESSAGE_WORD_01_BIT_1', class BC Messages, trigger "64_Message_Data_BC_MESSAGE_WORD_01" bit 9
   299: 'BC_MESSAGE_WORD_01_BIT_2', class BC Messages, trigger "64_Message_Data_BC_MESSAGE_WORD_01" bit 10
   295: 'BC_MESSAGE_WORD_01_BIT_14', class BC Messages, trigger "64_Message_Data_BC_MESSAGE_WORD_01" bit 6
   303: 'BC_MESSAGE_WORD_01_BIT_6', class BC Messages, trigger "64_Message_Data_BC_MESSAGE_WORD_01" bit 14
   301: 'BC_MESSAGE_WORD_01_BIT_4', class BC Messages, trigger "64_Message_Data_BC_MESSAGE_WORD_01" bit 12
   302: 'BC_MESSAGE_WORD_01_BIT_5', class BC Messages, trigger "64_Message_Data_BC_MESSAGE_WORD_01" bit 13
   310: 'BC_MESSAGE_WORD_02_BIT_13', class BC Messages, trigger "64_Message_Data_BC_MESSAGE_WORD_02" bit 5
   285: 'IGG_MESSAGE_WORD_02_BIT_4', class IGG Messages, trigger "64_Message_Data_IGG_MESSAGE_WORD_02" bit 12
   314: 'BC_MESSAGE_WORD_02_BIT_1', class BC Messages, trigger "64_Message_Data_BC_MESSAGE_WORD_02" bit 9
   287: 'IGG_MESSAGE_WORD_02_BIT_6', class IGG Messages, trigger "64_Message_Data_IGG_MESSAGE_WORD_02" bit 14